   1290: 'Carrier 20 Safe Output Card Fault', class No Acknowledgement, trigger "DB302_HMI_Faults_Carrier20_Faults_0" bit 9
   1291: 'Carrier 20 Standard Input Card Fault', class No Acknowledgement, trigger "DB302_HMI_Faults_Carrier20_Faults_0" bit 10
   1292: 'Carrier 20 Standard Output Card Fault', class No Acknowledgement, trigger "DB302_HMI_Faults_Carrier20_Faults_0" bit 11
   1293: 'Carrier 20 Encoder Position Fault', class No Acknowledgement, trigger "DB302_HMI_Faults_Carrier20_Faults_0" bit 12
   1294: 'Carrier 20 Encoder Internal Error', class No Acknowledgement, trigger "DB302_HMI_Faults_Carrier20_Faults_0" bit 13
   1295: 'Carrier 20 Encoder Comm Fault', class No Acknowledgement, trigger "DB302_HMI_Faults_Carrier20_Faults_0" bit 14
   1296: 'Carrier 20 HMI Comm Fault', class No Acknowledgement, trigger "DB302_HMI_Faults_Carrier20_Faults_0" bit 15
   1297: 'Carrier 20 Crash Detection Fault', class No Acknowledgement, trigger "DB302_HMI_Faults_Carrier20_Faults_1" bit 0
   1298: 'Carrier 20 Carrier Number Invalid', class No Acknowledgement, trigger "DB302_HMI_Faults_Carrier20_Faults_1" bit 1
   1299: 'Carrier 20 Drive: PROFINET configuration error', class No Acknowledgement, trigger "DB302_HMI_Faults_Carrier20_Faults_1" bit 2
   1300: 'Carrier 20 Drive: Error internal communications', class No Acknowledgement, trigger "DB302_HMI_Faults_Carrier20_Faults_1" bit 3
   1301: 'Carrier 20 Drive: Motor overtemperature', class No Acknowledgement, trigger "DB302_HMI_Faults_Carrier20_Faults_1" bit 4
   1302: 'Carrier 20 Drive: Motor overcurrent', class No Acknowledgement, trigger "DB302_HMI_Faults_Carrier20_Faults_1" bit 5
   1303: 'Carrier 20 Drive: Infeed or power unit not ready', class No Acknowledgement, trigger "DB302_HMI_Faults_Carrier20_Faults_1" bit 6
   1304: 'Carrier 20 Drive: Short-circuit/ground fault detected', class No Acknowledgement, trigger "DB302_HMI_Faults_Carrier20_Faults_1" bit 7
   1305: 'Carrier 20 Drive: PROFINET Setpoint timeout', class No Acknowledgement, trigger "DB302_HMI_Faults_Carrier20_Faults_1" bit 8
   1306: 'Carrier 20 Power unit: Overcurrent', class No Acknowledgement, trigger "DB302_HMI_Faults_Carrier20_Faults_1" bit 9
   1307: 'Carrier 20 Power unit: DC link voltage overvoltage', class No Acknowledgement, trigger "DB302_HMI_Faults_Carrier20_Faults_1" bit 10
   1308: 'Carrier 20 Power unit: DC link voltage undervoltage', class No Acknowledgement, trigger "DB302_HMI_Faults_Carrier20_Faults_1" bit 11
   1309: 'Carrier 20 Power unit: Line phase failure in main circuit', class No Acknowledgement, trigger "DB302_HMI_Faults_Carrier20_Faults_1" bit 12
   1310: 'Carrier 20 Power unit: Phase failure motor cable', class No Acknowledgement, trigger "DB302_HMI_Faults_Carrier20_Faults_1" bit 13
   1311: 'Carrier 20 Power unit: Ground fault', class No Acknowledgement, trigger "DB302_HMI_Faults_Carrier20_Faults_1" bit 14
   1312: 'Spare_Fault_1312', class No Acknowledgement, trigger "DB302_HMI_Faults_Carrier20_Faults_1" bit 15
   1313: 'Carrier 20 Motion Off Fault', class No Acknowledgement, trigger "DB302_HMI_Faults_Carrier20_Faults_2" bit 0
   1314: 'Carrier 20 Motion On Fault', class No Acknowledgement, trigger "DB302_HMI_Faults_Carrier20_Faults_2" bit 1
   1315: 'Carrier 20 Spacing Fault', class No Acknowledgement, trigger "DB302_HMI_Faults_Carrier20_Faults_2" bit 2
   1316: 'Carrier 20 Duplicate Carrier Number Fault', class No Acknowledgement, trigger "DB302_HMI_Faults_Carrier20_Faults_2" bit 3
   1317: 'Spare_Fault_1317', class No Acknowledgement, trigger "DB302_HMI_Faults_Carrier20_Faults_2" bit 4
   1318: 'Spare_Fault_1318', class No Acknowledgement, trigger "DB302_HMI_Faults_Carrier20_Faults_2" bit 5
   1319: 'Spare_Fault_1319', class No Acknowledgement, trigger "DB302_HMI_Faults_Carrier20_Faults_2" bit 6
   1320: 'Spare_Fault_1320', class No Acknowledgement, trigger "DB302_HMI_Faults_Carrier20_Faults_2" bit 7
   1321: 'Spare_Fault_1321', class No Acknowledgement, trigger "DB302_HMI_Faults_Carrier20_Faults_2" bit 8
   1322: 'Spare_Fault_1322', class No Acknowledgement, trigger "DB302_HMI_Faults_Carrier20_Faults_2" bit 9
   1323: 'Spare_Fault_1323', class No Acknowledgement, trigger "DB302_HMI_Faults_Carrier20_Faults_2" bit 10
   1324: 'Spare_Fault_1324', class No Acknowledgement, trigger "DB302_HMI_Faults_Carrier20_Faults_2" bit 11
   1325: 'Spare_Fault_1325', class No Acknowledgement, trigger "DB302_HMI_Faults_Carrier20_Faults_2" bit 12
   1326: 'Spare_Fault_1326', class No Acknowledgement, trigger "DB302_HMI_Faults_Carrier20_Faults_2" bit 13
   1327: 'Spare_Fault_1327', class No Acknowledgement, trigger "DB302_HMI_Faults_Carrier20_Faults_2" bit 14
   1328: 'Spare_Fault_1328', class No Acknowledgement, trigger "DB302_HMI_Faults_Carrier20_Faults_2" bit 15
   1329: 'Spare_Fault_1329', class No Acknowledgement, trigger "DB302_HMI_Faults_Carrier20_Faults_3" bit 0
   1330: 'Spare_Fault_1330', class No Acknowledgement, trigger "DB302_HMI_Faults_Carrier20_Faults_3" bit 1
   1331: 'Spare_Fault_1331', class No Acknowledgement, trigger "DB302_HMI_Faults_Carrier20_Faults_3" bit 2
   1332: 'Spare_Fault_1332', class No Acknowledgement, trigger "DB302_HMI_Faults_Carrier20_Faults_3" bit 3
   1333: 'Spare_Fault_1333', class No Acknowledgement, trigger "DB302_HMI_Faults_Carrier20_Faults_3" bit 4
   1334: 'Spare_Fault_1334', class No Acknowledgement, trigger "DB302_HMI_Faults_Carrier20_Faults_3" bit 5
   1335: 'Spare_Fault_1335', class No Acknowledgement, trigger "DB302_HMI_Faults_Carrier20_Faults_3" bit 6
   1336: 'Spare_Fault_1336', class No Acknowledgement, trigger "DB302_HMI_Faults_Carrier20_Faults_3" bit 7
   1337: 'Spare_Fault_1337', class No Acknowledgement, trigger "DB302_HMI_Faults_Carrier20_Faults_3" bit 8
   1338: 'Spare_Fault_1338', class No Acknowledgement, trigger "DB302_HMI_Faults_Carrier20_Faults_3" bit 9
   1339: 'Spare_Fault_1339', class No Acknowledgement, trigger "DB302_HMI_Faults_Carrier20_Faults_3" bit 10
   1340: 'Spare_Fault_1340', class No Acknowledgement, trigger "DB302_HMI_Faults_Carrier20_Faults_3" bit 11
   1341: 'Spare_Fault_1341', class No Acknowledgement, trigger "DB302_HMI_Faults_Carrier20_Faults_3" bit 12
   1342: 'Spare_Fault_1342', class No Acknowledgement, trigger "DB302_HMI_Faults_Carrier20_Faults_3" bit 13
   1343: 'Spare_Fault_1343', class No Acknowledgement, trigger "DB302_HMI_Faults_Carrier20_Faults_3" bit 14
   1344: 'Spare_Fault_1344', class No Acknowledgement, trigger "DB302_HMI_Faults_Carrier20_Faults_3" bit 15
   1345: 'Carrier 21 Disconnect Open Power Fault DI11.0', class No Acknowledgement, trigger "DB302_HMI_Faults_Carrier21_Faults_0" bit 0
   1346: 'Carrier 21 Drive Profinet Comm Fault', class No Acknowledgement, trigger "DB302_HMI_Faults_Carrier21_Faults_0" bit 1
   1347: 'Carrier 21 Production Stop Not Reset', class No Acknowledgement, trigger "DB302_HMI_Faults_Carrier21_Faults_0" bit 2
   1348: 'Carrier 21 CB02122 Tripped', class No Acknowledgement, trigger "DB302_HMI_Faults_Carrier21_Faults_0" bit 3
   1349: 'Carrier 21 CB02123 Tripped', class No Acknowledgement, trigger "DB302_HMI_Faults_Carrier21_Faults_0" bit 4
   1350: 'Carrier 21 AUX1 CB Tripped', class No Acknowledgement, trigger "DB302_HMI_Faults_Carrier21_Faults_0" bit 5
   1351: 'Carrier 21 AUX2 CB Tripped', class No Acknowledgement, trigger "DB302_HMI_Faults_Carrier21_Faults_0" bit 6
   1352: 'Carrier 21 PLC Not Communicating', class No Acknowledgement, trigger "DB302_HMI_Faults_Carrier21_Faults_0" bit 7
   1353: 'Carrier 21 Safe Input Card Fault', class No Acknowledgement, trigger "DB302_HMI_Faults_Carrier21_Faults_0" bit 8
   1354: 'Carrier 21 Safe Output Card Fault', class No Acknowledgement, trigger "DB302_HMI_Faults_Carrier21_Faults_0" bit 9
   1355: 'Carrier 21 Standard Input Card Fault', class No Acknowledgement, trigger "DB302_HMI_Faults_Carrier21_Faults_0" bit 10
   1356: 'Carrier 21 Standard Output Card Fault', class No Acknowledgement, trigger "DB302_HMI_Faults_Carrier21_Faults_0" bit 11
   1357: 'Carrier 21 Encoder Position Fault', class No Acknowledgement, trigger "DB302_HMI_Faults_Carrier21_Faults_0" bit 12
   1358: 'Carrier 21 Encoder Internal Error', class No Acknowledgement, trigger "DB302_HMI_Faults_Carrier21_Faults_0" bit 13
   1359: 'Carrier 21 Encoder Comm Fault', class No Acknowledgement, trigger "DB302_HMI_Faults_Carrier21_Faults_0" bit 14
   1360: 'Carrier 21 HMI Comm Fault', class No Acknowledgement, trigger "DB302_HMI_Faults_Carrier21_Faults_0" bit 15
   1361: 'Carrier 21 Crash Detection Fault', class No Acknowledgement, trigger "DB302_HMI_Faults_Carrier21_Faults_1" bit 0
   1362: 'Carrier 21 Carrier Number Invalid', class No Acknowledgement, trigger "DB302_HMI_Faults_Carrier21_Faults_1" bit 1
   1363: 'Carrier 21 Drive: PROFINET configuration error', class No Acknowledgement, trigger "DB302_HMI_Faults_Carrier21_Faults_1" bit 2
   1364: 'Carrier 21 Drive: Error internal communications', class No Acknowledgement, trigger "DB302_HMI_Faults_Carrier21_Faults_1" bit 3
   1365: 'Carrier 21 Drive: Motor overtemperature', class No Acknowledgement, trigger "DB302_HMI_Faults_Carrier21_Faults_1" bit 4
   1366: 'Carrier 21 Drive: Motor overcurrent', class No Acknowledgement, trigger "DB302_HMI_Faults_Carrier21_Faults_1" bit 5
   1367: 'Carrier 21 Drive: Infeed or power unit not ready', class No Acknowledgement, trigger "DB302_HMI_Faults_Carrier21_Faults_1" bit 6
   1368: 'Carrier 21 Drive: Short-circuit/ground fault detected', class No Acknowledgement, trigger "DB302_HMI_Faults_Carrier21_Faults_1" bit 7
   1369: 'Carrier 21 Drive: PROFINET Setpoint timeout', class No Acknowledgement, trigger "DB302_HMI_Faults_Carrier21_Faults_1" bit 8
   1370: 'Carrier 21 Power unit: Overcurrent', class No Acknowledgement, trigger "DB302_HMI_Faults_Carrier21_Faults_1" bit 9
   1371: 'Carrier 21 Power unit: DC link voltage overvoltage', class No Acknowledgement, trigger "DB302_HMI_Faults_Carrier21_Faults_1" bit 10
   1372: 'Carrier 21 Power unit: DC link voltage undervoltage', class No Acknowledgement, trigger "DB302_HMI_Faults_Carrier21_Faults_1" bit 11
   1373: 'Carrier 21 Power unit: Line phase failure in main circuit', class No Acknowledgement, trigger "DB302_HMI_Faults_Carrier21_Faults_1" bit 12
   1374: 'Carrier 21 Power unit: Phase failure motor cable', class No Acknowledgement, trigger "DB302_HMI_Faults_Carrier21_Faults_1" bit 13
   1375: 'Carrier 21 Power unit: Ground fault', class No Acknowledgement, trigger "DB302_HMI_Faults_Carrier21_Faults_1" bit 14
   1376: 'Spare_Fault_1376', class No Acknowledgement, trigger "DB302_HMI_Faults_Carrier21_Faults_1" bit 15
   1377: 'Carrier 21 Motion Off Fault', class No Acknowledgement, trigger "DB302_HMI_Faults_Carrier21_Faults_2" bit 0
   1378: 'Carrier 21 Motion On Fault', class No Acknowledgement, trigger "DB302_HMI_Faults_Carrier21_Faults_2" bit 1
   1379: 'Carrier 21 Spacing Fault', class No Acknowledgement, trigger "DB302_HMI_Faults_Carrier21_Faults_2" bit 2
   1380: 'Carrier 21 Duplicate Carrier Number Fault', class No Acknowledgement, trigger "DB302_HMI_Faults_Carrier21_Faults_2" bit 3
   1381: 'Spare_Fault_1381', class No Acknowledgement, trigger "DB302_HMI_Faults_Carrier21_Faults_2" bit 4
   1382: 'Spare_Fault_1382', class No Acknowledgement, trigger "DB302_HMI_Faults_Carrier21_Faults_2" bit 5
   1383: 'Spare_Fault_1383', class No Acknowledgement, trigger "DB302_HMI_Faults_Carrier21_Faults_2" bit 6
   1384: 'Spare_Fault_1384', class No Acknowledgement, trigger "DB302_HMI_Faults_Carrier21_Faults_2" bit 7
   1385: 'Spare_Fault_1385', class No Acknowledgement, trigger "DB302_HMI_Faults_Carrier21_Faults_2" bit 8
   1386: 'Spare_Fault_1386', class No Acknowledgement, trigger "DB302_HMI_Faults_Carrier21_Faults_2" bit 9
   1387: 'Spare_Fault_1387', class No Acknowledgement, trigger "DB302_HMI_Faults_Carrier21_Faults_2" bit 10
   1388: 'Spare_Fault_1388', class No Acknowledgement, trigger "DB302_HMI_Faults_Carrier21_Faults_2" bit 11
   1389: 'Spare_Fault_1389', class No Acknowledgement, trigger "DB302_HMI_Faults_Carrier21_Faults_2" bit 12
   1390: 'Spare_Fault_1390', class No Acknowledgement, trigger "DB302_HMI_Faults_Carrier21_Faults_2" bit 13
   1391: 'Spare_Fault_1391', class No Acknowledgement, trigger "DB302_HMI_Faults_Carrier21_Faults_2" bit 14
   1392: 'Spare_Fault_1392', class No Acknowledgement, trigger "DB302_HMI_Faults_Carrier21_Faults_2" bit 15
   1393: 'Spare_Fault_1393', class No Acknowledgement, trigger "DB302_HMI_Faults_Carrier21_Faults_3" bit 0
   1394: 'Spare_Fault_1394', class No Acknowledgement, trigger "DB302_HMI_Faults_Carrier21_Faults_3" bit 1
   1395: 'Spare_Fault_1395', class No Acknowledgement, trigger "DB302_HMI_Faults_Carrier21_Faults_3" bit 2
   1396: 'Spare_Fault_1396', class No Acknowledgement, trigger "DB302_HMI_Faults_Carrier21_Faults_3" bit 3
   1397: 'Spare_Fault_1397', class No Acknowledgement, trigger "DB302_HMI_Faults_Carrier21_Faults_3" bit 4
   1398: 'Spare_Fault_1398', class No Acknowledgement, trigger "DB302_HMI_Faults_Carrier21_Faults_3" bit 5
   1399: 'Spare_Fault_1399', class No Acknowledgement, trigger "DB302_HMI_Faults_Carrier21_Faults_3" bit 6
   1400: 'Spare_Fault_1400', class No Acknowledgement, trigger "DB302_HMI_Faults_Carrier21_Faults_3" bit 7
   1401: 'Spare_Fault_1401', class No Acknowledgement, trigger "DB302_HMI_Faults_Carrier21_Faults_3" bit 8
   1402: 'Spare_Fault_1402', class No Acknowledgement, trigger "DB302_HMI_Faults_Carrier21_Faults_3" bit 9
   1403: 'Spare_Fault_1403', class No Acknowledgement, trigger "DB302_HMI_Faults_Carrier21_Faults_3" bit 10
   1404: 'Spare_Fault_1404', class No Acknowledgement, trigger "DB302_HMI_Faults_Carrier21_Faults_3" bit 11
   1405: 'Spare_Fault_1405', class No Acknowledgement, trigger "DB302_HMI_Faults_Carrier21_Faults_3" bit 12
   1406: 'Spare_Fault_1406', class No Acknowledgement, trigger "DB302_HMI_Faults_Carrier21_Faults_3" bit 13
   1407: 'Spare_Fault_1407', class No Acknowledgement, trigger "DB302_HMI_Faults_Carrier21_Faults_3" bit 14
   1408: 'Spare_Fault_1408', class No Acknowledgement, trigger "DB302_HMI_Faults_Carrier21_Faults_3" bit 15
   1409: 'Carrier 22 Disconnect Open Power Fault DI11.0', class No Acknowledgement, trigger "DB302_HMI_Faults_Carrier22_Faults_0" bit 0
   1410: 'Carrier 22 Drive Profinet Comm Fault', class No Acknowledgement, trigger "DB302_HMI_Faults_Carrier22_Faults_0" bit 1
   1411: 'Carrier 22 Production Stop Not Reset', class No Acknowledgement, trigger "DB302_HMI_Faults_Carrier22_Faults_0" bit 2
   1412: 'Carrier 22 CB02122 Tripped', class No Acknowledgement, trigger "DB302_HMI_Faults_Carrier22_Faults_0" bit 3
   1413: 'Carrier 22 CB02123 Tripped', class No Acknowledgement, trigger "DB302_HMI_Faults_Carrier22_Faults_0" bit 4
   1414: 'Carrier 22 AUX1 CB Tripped', class No Acknowledgement, trigger "DB302_HMI_Faults_Carrier22_Faults_0" bit 5
   1415: 'Carrier 22 AUX2 CB Tripped', class No Acknowledgement, trigger "DB302_HMI_Faults_Carrier22_Faults_0" bit 6
   1416: 'Carrier 22 PLC Not Communicating', class No Acknowledgement, trigger "DB302_HMI_Faults_Carrier22_Faults_0" bit 7
   1417: 'Carrier 22 Safe Input Card Fault', class No Acknowledgement, trigger "DB302_HMI_Faults_Carrier22_Faults_0" bit 8
   1418: 'Carrier 22 Safe Output Card Fault', class No Acknowledgement, trigger "DB302_HMI_Faults_Carrier22_Faults_0" bit 9
   1419: 'Carrier 22 Standard Input Card Fault', class No Acknowledgement, trigger "DB302_HMI_Faults_Carrier22_Faults_0" bit 10
   1420: 'Carrier 22 Standard Output Card Fault', class No Acknowledgement, trigger "DB302_HMI_Faults_Carrier22_Faults_0" bit 11
   1421: 'Carrier 22 Encoder Position Fault', class No Acknowledgement, trigger "DB302_HMI_Faults_Carrier22_Faults_0" bit 12
   1422: 'Carrier 22 Encoder Internal Error', class No Acknowledgement, trigger "DB302_HMI_Faults_Carrier22_Faults_0" bit 13
   1423: 'Carrier 22 Encoder Comm Fault', class No Acknowledgement, trigger "DB302_HMI_Faults_Carrier22_Faults_0" bit 14
   1424: 'Carrier 22 HMI Comm Fault', class No Acknowledgement, trigger "DB302_HMI_Faults_Carrier22_Faults_0" bit 15
   1425: 'Carrier 22 Crash Detection Fault', class No Acknowledgement, trigger "DB302_HMI_Faults_Carrier22_Faults_1" bit 0
   1426: 'Carrier 22 Carrier Number Invalid', class No Acknowledgement, trigger "DB302_HMI_Faults_Carrier22_Faults_1" bit 1
   1427: 'Carrier 22 Drive: PROFINET configuration error', class No Acknowledgement, trigger "DB302_HMI_Faults_Carrier22_Faults_1" bit 2
   1428: 'Carrier 22 Drive: Error internal communications', class No Acknowledgement, trigger "DB302_HMI_Faults_Carrier22_Faults_1" bit 3
   1429: 'Carrier 22 Drive: Motor overtemperature', class No Acknowledgement, trigger "DB302_HMI_Faults_Carrier22_Faults_1" bit 4
   1430: 'Carrier 22 Drive: Motor overcurrent', class No Acknowledgement, trigger "DB302_HMI_Faults_Carrier22_Faults_1" bit 5
   1431: 'Carrier 22 Drive: Infeed or power unit not ready', class No Acknowledgement, trigger "DB302_HMI_Faults_Carrier22_Faults_1" bit 6
   1432: 'Carrier 22 Drive: Short-circuit/ground fault detected', class No Acknowledgement, trigger "DB302_HMI_Faults_Carrier22_Faults_1" bit 7
   1433: 'Carrier 22 Drive: PROFINET Setpoint timeout', class No Acknowledgement, trigger "DB302_HMI_Faults_Carrier22_Faults_1" bit 8
   1434: 'Carrier 22 Power unit: Overcurrent', class No Acknowledgement, trigger "DB302_HMI_Faults_Carrier22_Faults_1" bit 9
   1435: 'Carrier 22 Power unit: DC link voltage overvoltage', class No Acknowledgement, trigger "DB302_HMI_Faults_Carrier22_Faults_1" bit 10
   1436: 'Carrier 22 Power unit: DC link voltage undervoltage', class No Acknowledgement, trigger "DB302_HMI_Faults_Carrier22_Faults_1" bit 11
   1437: 'Carrier 22 Power unit: Line phase failure in main circuit', class No Acknowledgement, trigger "DB302_HMI_Faults_Carrier22_Faults_1" bit 12
   1438: 'Carrier 22 Power unit: Phase failure motor cable', class No Acknowledgement, trigger "DB302_HMI_Faults_Carrier22_Faults_1" bit 13
   1439: 'Carrier 22 Power unit: Ground fault', class No Acknowledgement, trigger "DB302_HMI_Faults_Carrier22_Faults_1" bit 14
   1440: 'Spare_Fault_1440', class No Acknowledgement, trigger "DB302_HMI_Faults_Carrier22_Faults_1" bit 15
   1441: 'Carrier 22 Motion Off Fault', class No Acknowledgement, trigger "DB302_HMI_Faults_Carrier22_Faults_2" bit 0
   1442: 'Carrier 22 Motion On Fault', class No Acknowledgement, trigger "DB302_HMI_Faults_Carrier22_Faults_2" bit 1
   1443: 'Carrier 22 Spacing Fault', class No Acknowledgement, trigger "DB302_HMI_Faults_Carrier22_Faults_2" bit 2
   1444: 'Carrier 22 Duplicate Carrier Number Fault', class No Acknowledgement, trigger "DB302_HMI_Faults_Carrier22_Faults_2" bit 3
   1445: 'Spare_Fault_1445', class No Acknowledgement, trigger "DB302_HMI_Faults_Carrier22_Faults_2" bit 4
   1446: 'Spare_Fault_1446', class No Acknowledgement, trigger "DB302_HMI_Faults_Carrier22_Faults_2" bit 5
   1447: 'Spare_Fault_1447', class No Acknowledgement, trigger "DB302_HMI_Faults_Carrier22_Faults_2" bit 6
   1448: 'Spare_Fault_1448', class No Acknowledgement, trigger "DB302_HMI_Faults_Carrier22_Faults_2" bit 7
   1449: 'Spare_Fault_1449', class No Acknowledgement, trigger "DB302_HMI_Faults_Carrier22_Faults_2" bit 8
   1450: 'Spare_Fault_1450', class No Acknowledgement, trigger "DB302_HMI_Faults_Carrier22_Faults_2" bit 9
   1451: 'Spare_Fault_1451', class No Acknowledgement, trigger "DB302_HMI_Faults_Carrier22_Faults_2" bit 10
   1452: 'Spare_Fault_1452', class No Acknowledgement, trigger "DB302_HMI_Faults_Carrier22_Faults_2" bit 11
   1453: 'Spare_Fault_1453', class No Acknowledgement, trigger "DB302_HMI_Faults_Carrier22_Faults_2" bit 12
   1454: 'Spare_Fault_1454', class No Acknowledgement, trigger "DB302_HMI_Faults_Carrier22_Faults_2" bit 13
   1455: 'Spare_Fault_1455', class No Acknowledgement, trigger "DB302_HMI_Faults_Carrier22_Faults_2" bit 14
   1456: 'Spare_Fault_1456', class No Acknowledgement, trigger "DB302_HMI_Faults_Carrier22_Faults_2" bit 15
   1457: 'Spare_Fault_1457', class No Acknowledgement, trigger "DB302_HMI_Faults_Carrier22_Faults_3" bit 0
   1458: 'Spare_Fault_1458', class No Acknowledgement, trigger "DB302_HMI_Faults_Carrier22_Faults_3" bit 1
   1459: 'Spare_Fault_1459', class No Acknowledgement, trigger "DB302_HMI_Faults_Carrier22_Faults_3" bit 2
   1460: 'Spare_Fault_1460', class No Acknowledgement, trigger "DB302_HMI_Faults_Carrier22_Faults_3" bit 3
   1461: 'Spare_Fault_1461', class No Acknowledgement, trigger "DB302_HMI_Faults_Carrier22_Faults_3" bit 4
   1462: 'Spare_Fault_1462', class No Acknowledgement, trigger "DB302_HMI_Faults_Carrier22_Faults_3" bit 5
   1463: 'Spare_Fault_1463', class No Acknowledgement, trigger "DB302_HMI_Faults_Carrier22_Faults_3" bit 6
   1464: 'Spare_Fault_1464', class No Acknowledgement, trigger "DB302_HMI_Faults_Carrier22_Faults_3" bit 7
   1465: 'Spare_Fault_1465', class No Acknowledgement, trigger "DB302_HMI_Faults_Carrier22_Faults_3" bit 8
   1466: 'Spare_Fault_1466', class No Acknowledgement, trigger "DB302_HMI_Faults_Carrier22_Faults_3" bit 9
   1467: 'Spare_Fault_1467', class No Acknowledgement, trigger "DB302_HMI_Faults_Carrier22_Faults_3" bit 10
   1468: 'Spare_Fault_1468', class No Acknowledgement, trigger "DB302_HMI_Faults_Carrier22_Faults_3" bit 11
   1469: 'Spare_Fault_1469', class No Acknowledgement, trigger "DB302_HMI_Faults_Carrier22_Faults_3" bit 12
   1470: 'Spare_Fault_1470', class No Acknowledgement, trigger "DB302_HMI_Faults_Carrier22_Faults_3" bit 13
   1471: 'Spare_Fault_1471', class No Acknowledgement, trigger "DB302_HMI_Faults_Carrier22_Faults_3" bit 14
   1472: 'Spare_Fault_1472', class No Acknowledgement, trigger "DB302_HMI_Faults_Carrier22_Faults_3" bit 15
   1473: 'Carrier 23 Disconnect Open Power Fault DI11.0', class No Acknowledgement, trigger "DB302_HMI_Faults_Carrier23_Faults_0" bit 0
   1474: 'Carrier 23 Drive Profinet Comm Fault', class No Acknowledgement, trigger "DB302_HMI_Faults_Carrier23_Faults_0" bit 1
   1475: 'Carrier 23 Production Stop Not Reset', class No Acknowledgement, trigger "DB302_HMI_Faults_Carrier23_Faults_0" bit 2
   1476: 'Carrier 23 CB02122 Tripped', class No Acknowledgement, trigger "DB302_HMI_Faults_Carrier23_Faults_0" bit 3
   1477: 'Carrier 23 CB02123 Tripped', class No Acknowledgement, trigger "DB302_HMI_Faults_Carrier23_Faults_0" bit 4
   1478: 'Carrier 23 AUX1 CB Tripped', class No Acknowledgement, trigger "DB302_HMI_Faults_Carrier23_Faults_0" bit 5
   1479: 'Carrier 23 AUX2 CB Tripped', class No Acknowledgement, trigger "DB302_HMI_Faults_Carrier23_Faults_0" bit 6
   1480: 'Carrier 23 PLC Not Communicating', class No Acknowledgement, trigger "DB302_HMI_Faults_Carrier23_Faults_0" bit 7
   1481: 'Carrier 23 Safe Input Card Fault', class No Acknowledgement, trigger "DB302_HMI_Faults_Carrier23_Faults_0" bit 8
   1482: 'Carrier 23 Safe Output Card Fault', class No Acknowledgement, trigger "DB302_HMI_Faults_Carrier23_Faults_0" bit 9
   1483: 'Carrier 23 Standard Input Card Fault', class No Acknowledgement, trigger "DB302_HMI_Faults_Carrier23_Faults_0" bit 10
   1484: 'Carrier 23 Standard Output Card Fault', class No Acknowledgement, trigger "DB302_HMI_Faults_Carrier23_Faults_0" bit 11
   1485: 'Carrier 23 Encoder Position Fault', class No Acknowledgement, trigger "DB302_HMI_Faults_Carrier23_Faults_0" bit 12
   1486: 'Carrier 23 Encoder Internal Error', class No Acknowledgement, trigger "DB302_HMI_Faults_Carrier23_Faults_0" bit 13
   1487: 'Carrier 23 Encoder Comm Fault', class No Acknowledgement, trigger "DB302_HMI_Faults_Carrier23_Faults_0" bit 14
   1488: 'Carrier 23 HMI Comm Fault', class No Acknowledgement, trigger "DB302_HMI_Faults_Carrier23_Faults_0" bit 15
   1489: 'Carrier 23 Crash Detection Fault', class No Acknowledgement, trigger "DB302_HMI_Faults_Carrier23_Faults_1" bit 0
   1490: 'Carrier 23 Carrier Number Invalid', class No Acknowledgement, trigger "DB302_HMI_Faults_Carrier23_Faults_1" bit 1
   1491: 'Carrier 23 Drive: PROFINET configuration error', class No Acknowledgement, trigger "DB302_HMI_Faults_Carrier23_Faults_1" bit 2
   1492: 'Carrier 23 Drive: Error internal communications', class No Acknowledgement, trigger "DB302_HMI_Faults_Carrier23_Faults_1" bit 3
   1493: 'Carrier 23 Drive: Motor overtemperature', class No Acknowledgement, trigger "DB302_HMI_Faults_Carrier23_Faults_1" bit 4
   1494: 'Carrier 23 Drive: Motor overcurrent', class No Acknowledgement, trigger "DB302_HMI_Faults_Carrier23_Faults_1" bit 5
   1495: 'Carrier 23 Drive: Infeed or power unit not ready', class No Acknowledgement, trigger "DB302_HMI_Faults_Carrier23_Faults_1" bit 6
   1496: 'Carrier 23 Drive: Short-circuit/ground fault detected', class No Acknowledgement, trigger "DB302_HMI_Faults_Carrier23_Faults_1" bit 7
   1497: 'Carrier 23 Drive: PROFINET Setpoint timeout', class No Acknowledgement, trigger "DB302_HMI_Faults_Carrier23_Faults_1" bit 8
   1498: 'Carrier 23 Power unit: Overcurrent', class No Acknowledgement, trigger "DB302_HMI_Faults_Carrier23_Faults_1" bit 9
   1499: 'Carrier 23 Power unit: DC link voltage overvoltage', class No Acknowledgement, trigger "DB302_HMI_Faults_Carrier23_Faults_1" bit 10
   1500: 'Carrier 23 Power unit: DC link voltage undervoltage', class No Acknowledgement, trigger "DB302_HMI_Faults_Carrier23_Faults_1" bit 11
   1501: 'Carrier 23 Power unit: Line phase failure in main circuit', class No Acknowledgement, trigger "DB302_HMI_Faults_Carrier23_Faults_1" bit 12
   1502: 'Carrier 23 Power unit: Phase failure motor cable', class No Acknowledgement, trigger "DB302_HMI_Faults_Carrier23_Faults_1" bit 13
   1503: 'Carrier 23 Power unit: Ground fault', class No Acknowledgement, trigger "DB302_HMI_Faults_Carrier23_Faults_1" bit 14
   1504: 'Spare_Fault_1504', class No Acknowledgement, trigger "DB302_HMI_Faults_Carrier23_Faults_1" bit 15
   1505: 'Carrier 23 Motion Off Fault', class No Acknowledgement, trigger "DB302_HMI_Faults_Carrier23_Faults_2" bit 0
   1506: 'Carrier 23 Motion On Fault', class No Acknowledgement, trigger "DB302_HMI_Faults_Carrier23_Faults_2" bit 1
   1507: 'Carrier 23 Spacing Fault', class No Acknowledgement, trigger "DB302_HMI_Faults_Carrier23_Faults_2" bit 2
   1508: 'Carrier 23 Duplicate Carrier Number Fault', class No Acknowledgement, trigger "DB302_HMI_Faults_Carrier23_Faults_2" bit 3
   1509: 'Spare_Fault_1509', class No Acknowledgement, trigger "DB302_HMI_Faults_Carrier23_Faults_2" bit 4
   1510: 'Spare_Fault_1510', class No Acknowledgement, trigger "DB302_HMI_Faults_Carrier23_Faults_2" bit 5
   1511: 'Spare_Fault_1511', class No Acknowledgement, trigger "DB302_HMI_Faults_Carrier23_Faults_2" bit 6
   1512: 'Spare_Fault_1512', class No Acknowledgement, trigger "DB302_HMI_Faults_Carrier23_Faults_2" bit 7
   1513: 'Spare_Fault_1513', class No Acknowledgement, trigger "DB302_HMI_Faults_Carrier23_Faults_2" bit 8
   1514: 'Spare_Fault_1514', class No Acknowledgement, trigger "DB302_HMI_Faults_Carrier23_Faults_2" bit 9
   1515: 'Spare_Fault_1515', class No Acknowledgement, trigger "DB302_HMI_Faults_Carrier23_Faults_2" bit 10
   1516: 'Spare_Fault_1516', class No Acknowledgement, trigger "DB302_HMI_Faults_Carrier23_Faults_2" bit 11
   1517: 'Spare_Fault_1517', class No Acknowledgement, trigger "DB302_HMI_Faults_Carrier23_Faults_2" bit 12
   1518: 'Spare_Fault_1518', class No Acknowledgement, trigger "DB302_HMI_Faults_Carrier23_Faults_2" bit 13
   1519: 'Spare_Fault_1519', class No Acknowledgement, trigger "DB302_HMI_Faults_Carrier23_Faults_2" bit 14
   1520: 'Spare_Fault_1520', class No Acknowledgement, trigger "DB302_HMI_Faults_Carrier23_Faults_2" bit 15
   1521: 'Spare_Fault_1521', class No Acknowledgement, trigger "DB302_HMI_Faults_Carrier23_Faults_3" bit 0
   1522: 'Spare_Fault_1522', class No Acknowledgement, trigger "DB302_HMI_Faults_Carrier23_Faults_3" bit 1
   1523: 'Spare_Fault_1523', class No Acknowledgement, trigger "DB302_HMI_Faults_Carrier23_Faults_3" bit 2
   1524: 'Spare_Fault_1524', class No Acknowledgement, trigger "DB302_HMI_Faults_Carrier23_Faults_3" bit 3
   1525: 'Spare_Fault_1525', class No Acknowledgement, trigger "DB302_HMI_Faults_Carrier23_Faults_3" bit 4
   1526: 'Spare_Fault_1526', class No Acknowledgement, trigger "DB302_HMI_Faults_Carrier23_Faults_3" bit 5
   1527: 'Spare_Fault_1527', class No Acknowledgement, trigger "DB302_HMI_Faults_Carrier23_Faults_3" bit 6
   1528: 'Spare_Fault_1528', class No Acknowledgement, trigger "DB302_HMI_Faults_Carrier23_Faults_3" bit 7
   1529: 'Spare_Fault_1529', class No Acknowledgement, trigger "DB302_HMI_Faults_Carrier23_Faults_3" bit 8
   1530: 'Spare_Fault_1530', class No Acknowledgement, trigger "DB302_HMI_Faults_Carrier23_Faults_3" bit 9
   1531: 'Spare_Fault_1531', class No Acknowledgement, trigger "DB302_HMI_Faults_Carrier23_Faults_3" bit 10
   1532: 'Spare_Fault_1532', class No Acknowledgement, trigger "DB302_HMI_Faults_Carrier23_Faults_3" bit 11
   1533: 'Spare_Fault_1533', class No Acknowledgement, trigger "DB302_HMI_Faults_Carrier23_Faults_3" bit 12
   1534: 'Spare_Fault_1534', class No Acknowledgement, trigger "DB302_HMI_Faults_Carrier23_Faults_3" bit 13
   1535: 'Spare_Fault_1535', class No Acknowledgement, trigger "DB302_HMI_Faults_Carrier23_Faults_3" bit 14
   1536: 'Spare_Fault_1536', class No Acknowledgement, trigger "DB302_HMI_Faults_Carrier23_Faults_3" bit 15
   1537: 'Carrier 24 Disconnect Open Power Fault DI11.0', class No Acknowledgement, trigger "DB302_HMI_Faults_Carrier24_Faults_0" bit 0
   1538: 'Carrier 24 Drive Profinet Comm Fault', class No Acknowledgement, trigger "DB302_HMI_Faults_Carrier24_Faults_0" bit 1
   1539: 'Carrier 24 Production Stop Not Reset', class No Acknowledgement, trigger "DB302_HMI_Faults_Carrier24_Faults_0" bit 2
   1540: 'Carrier 24 CB02122 Tripped', class No Acknowledgement, trigger "DB302_HMI_Faults_Carrier24_Faults_0" bit 3
   1541: 'Carrier 24 CB02123 Tripped', class No Acknowledgement, trigger "DB302_HMI_Faults_Carrier24_Faults_0" bit 4
   1542: 'Carrier 24 AUX1 CB Tripped', class No Acknowledgement, trigger "DB302_HMI_Faults_Carrier24_Faults_0" bit 5
   1543: 'Carrier 24 AUX2 CB Tripped', class No Acknowledgement, trigger "DB302_HMI_Faults_Carrier24_Faults_0" bit 6
   1544: 'Carrier 24 PLC Not Communicating', class No Acknowledgement, trigger "DB302_HMI_Faults_Carrier24_Faults_0" bit 7
   1545: 'Carrier 24 Safe Input Card Fault', class No Acknowledgement, trigger "DB302_HMI_Faults_Carrier24_Faults_0" bit 8
   1546: 'Carrier 24 Safe Output Card Fault', class No Acknowledgement, trigger "DB302_HMI_Faults_Carrier24_Faults_0" bit 9
   1547: 'Carrier 24 Standard Input Card Fault', class No Acknowledgement, trigger "DB302_HMI_Faults_Carrier24_Faults_0" bit 10
   1548: 'Carrier 24 Standard Output Card Fault', class No Acknowledgement, trigger "DB302_HMI_Faults_Carrier24_Faults_0" bit 11
   1549: 'Carrier 24 Encoder Position Fault', class No Acknowledgement, trigger "DB302_HMI_Faults_Carrier24_Faults_0" bit 12
   1550: 'Carrier 24 Encoder Internal Error', class No Acknowledgement, trigger "DB302_HMI_Faults_Carrier24_Faults_0" bit 13
   1551: 'Carrier 24 Encoder Comm Fault', class No Acknowledgement, trigger "DB302_HMI_Faults_Carrier24_Faults_0" bit 14
   1552: 'Carrier 24 HMI Comm Fault', class No Acknowledgement, trigger "DB302_HMI_Faults_Carrier24_Faults_0" bit 15
   1553: 'Carrier 24 Crash Detection Fault', class No Acknowledgement, trigger "DB302_HMI_Faults_Carrier24_Faults_1" bit 0
   1554: 'Carrier 24 Carrier Number Invalid', class No Acknowledgement, trigger "DB302_HMI_Faults_Carrier24_Faults_1" bit 1
   1555: 'Carrier 24 Drive: PROFINET configuration error', class No Acknowledgement, trigger "DB302_HMI_Faults_Carrier24_Faults_1" bit 2
   1556: 'Carrier 24 Drive: Error internal communications', class No Acknowledgement, trigger "DB302_HMI_Faults_Carrier24_Faults_1" bit 3
   1557: 'Carrier 24 Drive: Motor overtemperature', class No Acknowledgement, trigger "DB302_HMI_Faults_Carrier24_Faults_1" bit 4
   1558: 'Carrier 24 Drive: Motor overcurrent', class No Acknowledgement, trigger "DB302_HMI_Faults_Carrier24_Faults_1" bit 5
   1559: 'Carrier 24 Drive: Infeed or power unit not ready', class No Acknowledgement, trigger "DB302_HMI_Faults_Carrier24_Faults_1" bit 6
   1560: 'Carrier 24 Drive: Short-circuit/ground fault detected', class No Acknowledgement, trigger "DB302_HMI_Faults_Carrier24_Faults_1" bit 7
   1561: 'Carrier 24 Drive: PROFINET Setpoint timeout', class No Acknowledgement, trigger "DB302_HMI_Faults_Carrier24_Faults_1" bit 8
   1562: 'Carrier 24 Power unit: Overcurrent', class No Acknowledgement, trigger "DB302_HMI_Faults_Carrier24_Faults_1" bit 9
   1563: 'Carrier 24 Power unit: DC link voltage overvoltage', class No Acknowledgement, trigger "DB302_HMI_Faults_Carrier24_Faults_1" bit 10
   1564: 'Carrier 24 Power unit: DC link voltage undervoltage', class No Acknowledgement, trigger "DB302_HMI_Faults_Carrier24_Faults_1" bit 11
   1565: 'Carrier 24 Power unit: Line phase failure in main circuit', class No Acknowledgement, trigger "DB302_HMI_Faults_Carrier24_Faults_1" bit 12
   1566: 'Carrier 24 Power unit: Phase failure motor cable', class No Acknowledgement, trigger "DB302_HMI_Faults_Carrier24_Faults_1" bit 13
   1567: 'Carrier 24 Power unit: Ground fault', class No Acknowledgement, trigger "DB302_HMI_Faults_Carrier24_Faults_1" bit 14
   1568: 'Spare_Fault_1568', class No Acknowledgement, trigger "DB302_HMI_Faults_Carrier24_Faults_1" bit 15
   1569: 'Carrier 24 Motion Off Fault', class No Acknowledgement, trigger "DB302_HMI_Faults_Carrier24_Faults_2" bit 0
   1570: 'Carrier 24 Motion On Fault', class No Acknowledgement, trigger "DB302_HMI_Faults_Carrier24_Faults_2" bit 1
   1571: 'Carrier 24 Spacing Fault', class No Acknowledgement, trigger "DB302_HMI_Faults_Carrier24_Faults_2" bit 2
   1572: 'Carrier 24 Duplicate Carrier Number Fault', class No Acknowledgement, trigger "DB302_HMI_Faults_Carrier24_Faults_2" bit 3
   1573: 'Spare_Fault_1573', class No Acknowledgement, trigger "DB302_HMI_Faults_Carrier24_Faults_2" bit 4
   1574: 'Spare_Fault_1574', class No Acknowledgement, trigger "DB302_HMI_Faults_Carrier24_Faults_2" bit 5
   1575: 'Spare_Fault_1575', class No Acknowledgement, trigger "DB302_HMI_Faults_Carrier24_Faults_2" bit 6
   1576: 'Spare_Fault_1576', class No Acknowledgement, trigger "DB302_HMI_Faults_Carrier24_Faults_2" bit 7
   1577: 'Spare_Fault_1577', class No Acknowledgement, trigger "DB302_HMI_Faults_Carrier24_Faults_2" bit 8
   1578: 'Spare_Fault_1578', class No Acknowledgement, trigger "DB302_HMI_Faults_Carrier24_Faults_2" bit 9
   1579: 'Spare_Fault_1579', class No Acknowledgement, trigger "DB302_HMI_Faults_Carrier24_Faults_2" bit 10
   1580: 'Spare_Fault_1580', class No Acknowledgement, trigger "DB302_HMI_Faults_Carrier24_Faults_2" bit 11
   1581: 'Spare_Fault_1581', class No Acknowledgement, trigger "DB302_HMI_Faults_Carrier24_Faults_2" bit 12
   1582: 'Spare_Fault_1582', class No Acknowledgement, trigger "DB302_HMI_Faults_Carrier24_Faults_2" bit 13
   1583: 'Spare_Fault_1583', class No Acknowledgement, trigger "DB302_HMI_Faults_Carrier24_Faults_2" bit 14
   1584: 'Spare_Fault_1584', class No Acknowledgement, trigger "DB302_HMI_Faults_Carrier24_Faults_2" bit 15
   1585: 'Spare_Fault_1585', class No Acknowledgement, trigger "DB302_HMI_Faults_Carrier24_Faults_3" bit 0
   1586: 'Spare_Fault_1586', class No Acknowledgement, trigger "DB302_HMI_Faults_Carrier24_Faults_3" bit 1
   1587: 'Spare_Fault_1587', class No Acknowledgement, trigger "DB302_HMI_Faults_Carrier24_Faults_3" bit 2
   1588: 'Spare_Fault_1588', class No Acknowledgement, trigger "DB302_HMI_Faults_Carrier24_Faults_3" bit 3
   1589: 'Spare_Fault_1589', class No Acknowledgement, trigger "DB302_HMI_Faults_Carrier24_Faults_3" bit 4
   1590: 'Spare_Fault_1590', class No Acknowledgement, trigger "DB302_HMI_Faults_Carrier24_Faults_3" bit 5
   1591: 'Spare_Fault_1591', class No Acknowledgement, trigger "DB302_HMI_Faults_Carrier24_Faults_3" bit 6
   1592: 'Spare_Fault_1592', class No Acknowledgement, trigger "DB302_HMI_Faults_Carrier24_Faults_3" bit 7
   1593: 'Spare_Fault_1593', class No Acknowledgement, trigger "DB302_HMI_Faults_Carrier24_Faults_3" bit 8
   1594: 'Spare_Fault_1594', class No Acknowledgement, trigger "DB302_HMI_Faults_Carrier24_Faults_3" bit 9
   1595: 'Spare_Fault_1595', class No Acknowledgement, trigger "DB302_HMI_Faults_Carrier24_Faults_3" bit 10
   1596: 'Spare_Fault_1596', class No Acknowledgement, trigger "DB302_HMI_Faults_Carrier24_Faults_3" bit 11
   1597: 'Spare_Fault_1597', class No Acknowledgement, trigger "DB302_HMI_Faults_Carrier24_Faults_3" bit 12
   1598: 'Spare_Fault_1598', class No Acknowledgement, trigger "DB302_HMI_Faults_Carrier24_Faults_3" bit 13
   1599: 'Spare_Fault_1599', class No Acknowledgement, trigger "DB302_HMI_Faults_Carrier24_Faults_3" bit 14
   1600: 'Spare_Fault_1600', class No Acknowledgement, trigger "DB302_HMI_Faults_Carrier24_Faults_3" bit 15
   1601: 'Carrier 25 Disconnect Open Power Fault DI11.0', class No Acknowledgement, trigger "DB302_HMI_Faults_Carrier25_Faults_0" bit 0
   1602: 'Carrier 25 Drive Profinet Comm Fault', class No Acknowledgement, trigger "DB302_HMI_Faults_Carrier25_Faults_0" bit 1
   1603: 'Carrier 25 Production Stop Not Reset', class No Acknowledgement, trigger "DB302_HMI_Faults_Carrier25_Faults_0" bit 2
   1604: 'Carrier 25 CB02122 Tripped', class No Acknowledgement, trigger "DB302_HMI_Faults_Carrier25_Faults_0" bit 3
   1605: 'Carrier 25 CB02123 Tripped', class No Acknowledgement, trigger "DB302_HMI_Faults_Carrier25_Faults_0" bit 4
   1606: 'Carrier 25 AUX1 CB Tripped', class No Acknowledgement, trigger "DB302_HMI_Faults_Carrier25_Faults_0" bit 5
   1607: 'Carrier 25 AUX2 CB Tripped', class No Acknowledgement, trigger "DB302_HMI_Faults_Carrier25_Faults_0" bit 6
   1608: 'Carrier 25 PLC Not Communicating', class No Acknowledgement, trigger "DB302_HMI_Faults_Carrier25_Faults_0" bit 7
   1609: 'Carrier 25 Safe Input Card Fault', class No Acknowledgement, trigger "DB302_HMI_Faults_Carrier25_Faults_0" bit 8
   1610: 'Carrier 25 Safe Output Card Fault', class No Acknowledgement, trigger "DB302_HMI_Faults_Carrier25_Faults_0" bit 9
   1611: 'Carrier 25 Standard Input Card Fault', class No Acknowledgement, trigger "DB302_HMI_Faults_Carrier25_Faults_0" bit 10
   1612: 'Carrier 25 Standard Output Card Fault', class No Acknowledgement, trigger "DB302_HMI_Faults_Carrier25_Faults_0" bit 11
   1613: 'Carrier 25 Encoder Position Fault', class No Acknowledgement, trigger "DB302_HMI_Faults_Carrier25_Faults_0" bit 12
   1614: 'Carrier 25 Encoder Internal Error', class No Acknowledgement, trigger "DB302_HMI_Faults_Carrier25_Faults_0" bit 13
   1615: 'Carrier 25 Encoder Comm Fault', class No Acknowledgement, trigger "DB302_HMI_Faults_Carrier25_Faults_0" bit 14
   1616: 'Carrier 25 HMI Comm Fault', class No Acknowledgement, trigger "DB302_HMI_Faults_Carrier25_Faults_0" bit 15
   1617: 'Carrier 25 Crash Detection Fault', class No Acknowledgement, trigger "DB302_HMI_Faults_Carrier25_Faults_1" bit 0
   1618: 'Carrier 25 Carrier Number Invalid', class No Acknowledgement, trigger "DB302_HMI_Faults_Carrier25_Faults_1" bit 1
   1619: 'Carrier 25 Drive: PROFINET configuration error', class No Acknowledgement, trigger "DB302_HMI_Faults_Carrier25_Faults_1" bit 2
   1620: 'Carrier 25 Drive: Error internal communications', class No Acknowledgement, trigger "DB302_HMI_Faults_Carrier25_Faults_1" bit 3
   1621: 'Carrier 25 Drive: Motor overtemperature', class No Acknowledgement, trigger "DB302_HMI_Faults_Carrier25_Faults_1" bit 4
   1622: 'Carrier 25 Drive: Motor overcurrent', class No Acknowledgement, trigger "DB302_HMI_Faults_Carrier25_Faults_1" bit 5
   1623: 'Carrier 25 Drive: Infeed or power unit not ready', class No Acknowledgement, trigger "DB302_HMI_Faults_Carrier25_Faults_1" bit 6
   1624: 'Carrier 25 Drive: Short-circuit/ground fault detected', class No Acknowledgement, trigger "DB302_HMI_Faults_Carrier25_Faults_1" bit 7
   1625: 'Carrier 25 Drive: PROFINET Setpoint timeout', class No Acknowledgement, trigger "DB302_HMI_Faults_Carrier25_Faults_1" bit 8
   1626: 'Carrier 25 Power unit: Overcurrent', class No Acknowledgement, trigger "DB302_HMI_Faults_Carrier25_Faults_1" bit 9
   1627: 'Carrier 25 Power unit: DC link voltage overvoltage', class No Acknowledgement, trigger "DB302_HMI_Faults_Carrier25_Faults_1" bit 10
   1628: 'Carrier 25 Power unit: DC link voltage undervoltage', class No Acknowledgement, trigger "DB302_HMI_Faults_Carrier25_Faults_1" bit 11
   1629: 'Carrier 25 Power unit: Line phase failure in main circuit', class No Acknowledgement, trigger "DB302_HMI_Faults_Carrier25_Faults_1" bit 12
   1630: 'Carrier 25 Power unit: Phase failure motor cable', class No Acknowledgement, trigger "DB302_HMI_Faults_Carrier25_Faults_1" bit 13
   1631: 'Carrier 25 Power unit: Ground fault', class No Acknowledgement, trigger "DB302_HMI_Faults_Carrier25_Faults_1" bit 14
   1632: 'Spare_Fault_1632', class No Acknowledgement, trigger "DB302_HMI_Faults_Carrier25_Faults_1" bit 15
   1633: 'Carrier 25 Motion Off Fault', class No Acknowledgement, trigger "DB302_HMI_Faults_Carrier25_Faults_2" bit 0
   1634: 'Carrier 25 Motion On Fault', class No Acknowledgement, trigger "DB302_HMI_Faults_Carrier25_Faults_2" bit 1
   1635: 'Carrier 25 Spacing Fault', class No Acknowledgement, trigger "DB302_HMI_Faults_Carrier25_Faults_2" bit 2
   1636: 'Carrier 25 Duplicate Carrier Number Fault', class No Acknowledgement, trigger "DB302_HMI_Faults_Carrier25_Faults_2" bit 3
   1637: 'Spare_Fault_1637', class No Acknowledgement, trigger "DB302_HMI_Faults_Carrier25_Faults_2" bit 4
   1638: 'Spare_Fault_1638', class No Acknowledgement, trigger "DB302_HMI_Faults_Carrier25_Faults_2" bit 5
   1639: 'Spare_Fault_1639', class No Acknowledgement, trigger "DB302_HMI_Faults_Carrier25_Faults_2" bit 6
   1640: 'Spare_Fault_1640', class No Acknowledgement, trigger "DB302_HMI_Faults_Carrier25_Faults_2" bit 7
   1641: 'Spare_Fault_1641', class No Acknowledgement, trigger "DB302_HMI_Faults_Carrier25_Faults_2" bit 8
   1642: 'Spare_Fault_1642', class No Acknowledgement, trigger "DB302_HMI_Faults_Carrier25_Faults_2" bit 9
   1643: 'Spare_Fault_1643', class No Acknowledgement, trigger "DB302_HMI_Faults_Carrier25_Faults_2" bit 10
   1644: 'Spare_Fault_1644', class No Acknowledgement, trigger "DB302_HMI_Faults_Carrier25_Faults_2" bit 11
   1645: 'Spare_Fault_1645', class No Acknowledgement, trigger "DB302_HMI_Faults_Carrier25_Faults_2" bit 12
   1646: 'Spare_Fault_1646', class No Acknowledgement, trigger "DB302_HMI_Faults_Carrier25_Faults_2" bit 13
   1647: 'Spare_Fault_1647', class No Acknowledgement, trigger "DB302_HMI_Faults_Carrier25_Faults_2" bit 14
   1648: 'Spare_Fault_1648', class No Acknowledgement, trigger "DB302_HMI_Faults_Carrier25_Faults_2" bit 15
   1649: 'Spare_Fault_1649', class No Acknowledgement, trigger "DB302_HMI_Faults_Carrier25_Faults_3" bit 0
   1650: 'Spare_Fault_1650', class No Acknowledgement, trigger "DB302_HMI_Faults_Carrier25_Faults_3" bit 1
   1651: 'Spare_Fault_1651', class No Acknowledgement, trigger "DB302_HMI_Faults_Carrier25_Faults_3" bit 2
   1652: 'Spare_Fault_1652', class No Acknowledgement, trigger "DB302_HMI_Faults_Carrier25_Faults_3" bit 3
   1653: 'Spare_Fault_1653', class No Acknowledgement, trigger "DB302_HMI_Faults_Carrier25_Faults_3" bit 4
   1654: 'Spare_Fault_1654', class No Acknowledgement, trigger "DB302_HMI_Faults_Carrier25_Faults_3" bit 5
   1655: 'Spare_Fault_1655', class No Acknowledgement, trigger "DB302_HMI_Faults_Carrier25_Faults_3" bit 6
   1656: 'Spare_Fault_1656', class No Acknowledgement, trigger "DB302_HMI_Faults_Carrier25_Faults_3" bit 7
   1657: 'Spare_Fault_1657', class No Acknowledgement, trigger "DB302_HMI_Faults_Carrier25_Faults_3" bit 8
   1658: 'Spare_Fault_1658', class No Acknowledgement, trigger "DB302_HMI_Faults_Carrier25_Faults_3" bit 9
   1659: 'Spare_Fault_1659', class No Acknowledgement, trigger "DB302_HMI_Faults_Carrier25_Faults_3" bit 10
   1660: 'Spare_Fault_1660', class No Acknowledgement, trigger "DB302_HMI_Faults_Carrier25_Faults_3" bit 11
   1661: 'Spare_Fault_1661', class No Acknowledgement, trigger "DB302_HMI_Faults_Carrier25_Faults_3" bit 12
   1662: 'Spare_Fault_1662', class No Acknowledgement, trigger "DB302_HMI_Faults_Carrier25_Faults_3" bit 13
   1663: 'Spare_Fault_1663', class No Acknowledgement, trigger "DB302_HMI_Faults_Carrier25_Faults_3" bit 14
   1664: 'Spare_Fault_1664', class No Acknowledgement, trigger "DB302_HMI_Faults_Carrier25_Faults_3" bit 15
   1665: 'Carrier 26 Disconnect Open Power Fault DI11.0', class No Acknowledgement, trigger "DB302_HMI_Faults_Carrier26_Faults_0" bit 0
   1666: 'Carrier 26 Drive Profinet Comm Fault', class No Acknowledgement, trigger "DB302_HMI_Faults_Carrier26_Faults_0" bit 1
   1667: 'Carrier 26 Production Stop Not Reset', class No Acknowledgement, trigger "DB302_HMI_Faults_Carrier26_Faults_0" bit 2
   1668: 'Carrier 26 CB02122 Tripped', class No Acknowledgement, trigger "DB302_HMI_Faults_Carrier26_Faults_0" bit 3
   1669: 'Carrier 26 CB02123 Tripped', class No Acknowledgement, trigger "DB302_HMI_Faults_Carrier26_Faults_0" bit 4
   1670: 'Carrier 26 AUX1 CB Tripped', class No Acknowledgement, trigger "DB302_HMI_Faults_Carrier26_Faults_0" bit 5
   1671: 'Carrier 26 AUX2 CB Tripped', class No Acknowledgement, trigger "DB302_HMI_Faults_Carrier26_Faults_0" bit 6
   1672: 'Carrier 26 PLC Not Communicating', class No Acknowledgement, trigger "DB302_HMI_Faults_Carrier26_Faults_0" bit 7
   1673: 'Carrier 26 Safe Input Card Fault', class No Acknowledgement, trigger "DB302_HMI_Faults_Carrier26_Faults_0" bit 8
   1674: 'Carrier 26 Safe Output Card Fault', class No Acknowledgement, trigger "DB302_HMI_Faults_Carrier26_Faults_0" bit 9
   1675: 'Carrier 26 Standard Input Card Fault', class No Acknowledgement, trigger "DB302_HMI_Faults_Carrier26_Faults_0" bit 10
   1676: 'Carrier 26 Standard Output Card Fault', class No Acknowledgement, trigger "DB302_HMI_Faults_Carrier26_Faults_0" bit 11
   1677: 'Carrier 26 Encoder Position Fault', class No Acknowledgement, trigger "DB302_HMI_Faults_Carrier26_Faults_0" bit 12
   1678: 'Carrier 26 Encoder Internal Error', class No Acknowledgement, trigger "DB302_HMI_Faults_Carrier26_Faults_0" bit 13
   1679: 'Carrier 26 Encoder Comm Fault', class No Acknowledgement, trigger "DB302_HMI_Faults_Carrier26_Faults_0" bit 14
   1680: 'Carrier 26 HMI Comm Fault', class No Acknowledgement, trigger "DB302_HMI_Faults_Carrier26_Faults_0" bit 15
   1681: 'Carrier 26 Crash Detection Fault', class No Acknowledgement, trigger "DB302_HMI_Faults_Carrier26_Faults_1" bit 0
   1682: 'Carrier 26 Carrier Number Invalid', class No Acknowledgement, trigger "DB302_HMI_Faults_Carrier26_Faults_1" bit 1
   1683: 'Carrier 26 Drive: PROFINET configuration error', class No Acknowledgement, trigger "DB302_HMI_Faults_Carrier26_Faults_1" bit 2
   1684: 'Carrier 26 Drive: Error internal communications', class No Acknowledgement, trigger "DB302_HMI_Faults_Carrier26_Faults_1" bit 3
   1685: 'Carrier 26 Drive: Motor overtemperature', class No Acknowledgement, trigger "DB302_HMI_Faults_Carrier26_Faults_1" bit 4
   1686: 'Carrier 26 Drive: Motor overcurrent', class No Acknowledgement, trigger "DB302_HMI_Faults_Carrier26_Faults_1" bit 5
   1687: 'Carrier 26 Drive: Infeed or power unit not ready', class No Acknowledgement, trigger "DB302_HMI_Faults_Carrier26_Faults_1" bit 6
   1688: 'Carrier 26 Drive: Short-circuit/ground fault detected', class No Acknowledgement, trigger "DB302_HMI_Faults_Carrier26_Faults_1" bit 7
   1689: 'Carrier 26 Drive: PROFINET Setpoint timeout', class No Acknowledgement, trigger "DB302_HMI_Faults_Carrier26_Faults_1" bit 8
   1690: 'Carrier 26 Power unit: Overcurrent', class No Acknowledgement, trigger "DB302_HMI_Faults_Carrier26_Faults_1" bit 9
   1691: 'Carrier 26 Power unit: DC link voltage overvoltage', class No Acknowledgement, trigger "DB302_HMI_Faults_Carrier26_Faults_1" bit 10
   1692: 'Carrier 26 Power unit: DC link voltage undervoltage', class No Acknowledgement, trigger "DB302_HMI_Faults_Carrier26_Faults_1" bit 11
   1693: 'Carrier 26 Power unit: Line phase failure in main circuit', class No Acknowledgement, trigger "DB302_HMI_Faults_Carrier26_Faults_1" bit 12
   1694: 'Carrier 26 Power unit: Phase failure motor cable', class No Acknowledgement, trigger "DB302_HMI_Faults_Carrier26_Faults_1" bit 13
   1695: 'Carrier 26 Power unit: Ground fault', class No Acknowledgement, trigger "DB302_HMI_Faults_Carrier26_Faults_1" bit 14
   1696: 'Spare_Fault_1696', class No Acknowledgement, trigger "DB302_HMI_Faults_Carrier26_Faults_1" bit 15
   1697: 'Carrier 26 Motion Off Fault', class No Acknowledgement, trigger "DB302_HMI_Faults_Carrier26_Faults_2" bit 0
   1698: 'Carrier 26 Motion On Fault', class No Acknowledgement, trigger "DB302_HMI_Faults_Carrier26_Faults_2" bit 1
   1699: 'Carrier 26 Spacing Fault', class No Acknowledgement, trigger "DB302_HMI_Faults_Carrier26_Faults_2" bit 2
   1700: 'Carrier 26 Duplicate Carrier Number Fault', class No Acknowledgement, trigger "DB302_HMI_Faults_Carrier26_Faults_2" bit 3
   1701: 'Spare_Fault_1701', class No Acknowledgement, trigger "DB302_HMI_Faults_Carrier26_Faults_2" bit 4
   1702: 'Spare_Fault_1702', class No Acknowledgement, trigger "DB302_HMI_Faults_Carrier26_Faults_2" bit 5
   1703: 'Spare_Fault_1703', class No Acknowledgement, trigger "DB302_HMI_Faults_Carrier26_Faults_2" bit 6
   1704: 'Spare_Fault_1704', class No Acknowledgement, trigger "DB302_HMI_Faults_Carrier26_Faults_2" bit 7
   1705: 'Spare_Fault_1705', class No Acknowledgement, trigger "DB302_HMI_Faults_Carrier26_Faults_2" bit 8
   1706: 'Spare_Fault_1706', class No Acknowledgement, trigger "DB302_HMI_Faults_Carrier26_Faults_2" bit 9
   1707: 'Spare_Fault_1707', class No Acknowledgement, trigger "DB302_HMI_Faults_Carrier26_Faults_2" bit 10
   1708: 'Spare_Fault_1708', class No Acknowledgement, trigger "DB302_HMI_Faults_Carrier26_Faults_2" bit 11
